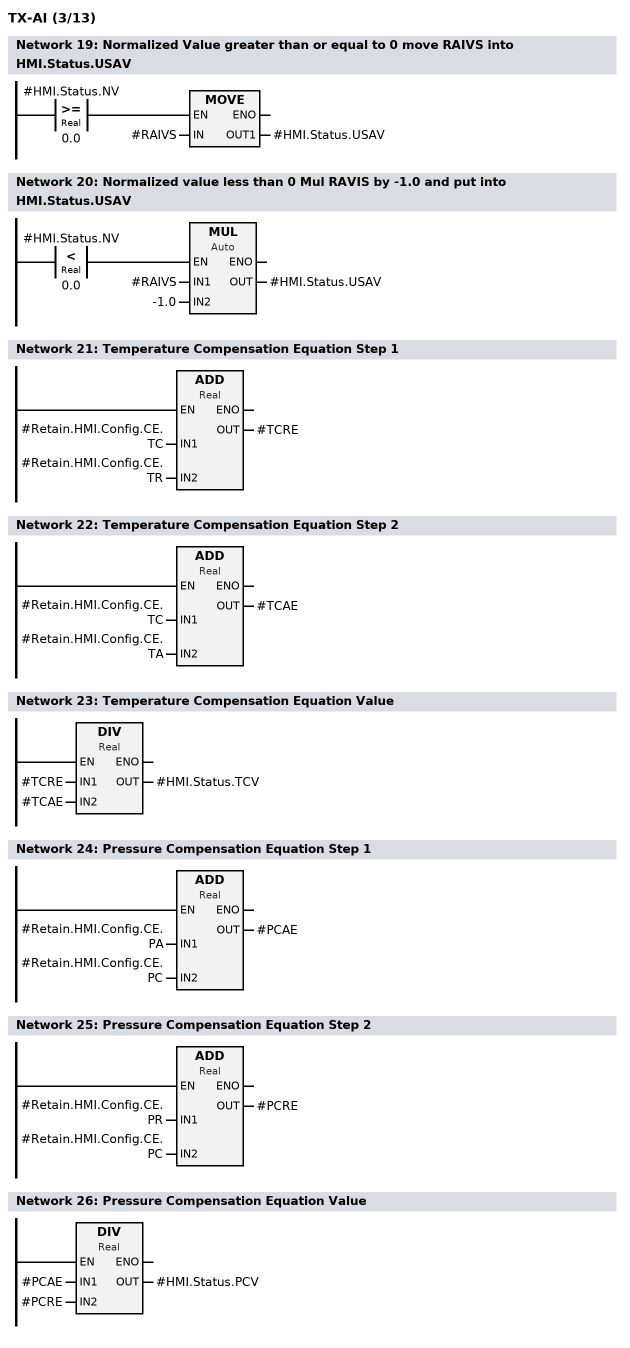
   RUNG wire#powerrail
      { S7_Templates := "SrcType := Real" } GE_Contact(in1 := #HMI.Status.NV, in2 := 0.0)
      { S7_GenerateENO := "TRUE" } Move(in := #RAIVS, out1 => #HMI.Status.USAV)
   END_RUNG
   // the same network as SCL:
   IF #HMI.Status.NV >= 0.0 THEN #HMI.Status.USAV := #RAIVS; END_IF;
END_REGION

REGION Network 20: Normalized value less than 0 Mul RAVIS by -1.0 and put into HMI.Status.USAV
   RUNG wire#powerrail
      { S7_Templates := "SrcType := Real" } LT_Contact(in1 := #HMI.Status.NV, in2 := 0.0)
      { S7_GenerateENO := "TRUE" } Mul(in1 := #RAIVS, in2 := -1.0, out => #HMI.Status.USAV)
   END_RUNG
   // the same network as SCL:
   IF #HMI.Status.NV < 0.0 THEN #HMI.Status.USAV := #RAIVS * (-1.0); END_IF;
END_REGION

REGION Network 21: Temperature Compensation Equation Step 1
   RUNG wire#powerrail
      { S7_Templates := "SrcType := Real"; S7_GenerateENO := "TRUE" } Add(in1 := #Retain.HMI.Config.CE.TC, in2 := #Retain.HMI.Config.CE.TR, out => #TCRE)
   END_RUNG
   // the same network as SCL:
   #TCRE := #Retain.HMI.Config.CE.TC + #Retain.HMI.Config.CE.TR;
END_REGION

REGION Network 22: Temperature Compensation Equation Step 2
   RUNG wire#powerrail
      { S7_Templates := "SrcType := Real"; S7_GenerateENO := "TRUE" } Add(in1 := #Retain.HMI.Config.CE.TC, in2 := #Retain.HMI.Config.CE.TA, out => #TCAE)
   END_RUNG
   // the same network as SCL:
   #TCAE := #Retain.HMI.Config.CE.TC + #Retain.HMI.Config.CE.TA;
END_REGION

REGION Network 23: Temperature Compensation Equation Value
   RUNG wire#powerrail
      { S7_Templates := "SrcType := Real"; S7_GenerateENO := "TRUE" } Div(in1 := #TCRE, in2 := #TCAE, out => #HMI.Status.TCV)
   END_RUNG
   // the same network as SCL:
   #HMI.Status.TCV := #TCRE / #TCAE;
END_REGION

REGION Network 24: Pressure Compensation Equation Step 1
   RUNG wire#powerrail
      { S7_Templates := "SrcType := Real"; S7_GenerateENO := "TRUE" } Add(in1 := #Retain.HMI.Config.CE.PA, in2 := #Retain.HMI.Config.CE.PC, out => #PCAE)
   END_RUNG
   // the same network as SCL:
   #PCAE := #Retain.HMI.Config.CE.PA + #Retain.HMI.Config.CE.PC;
END_REGION

REGION Network 25: Pressure Compensation Equation Step 2
   RUNG wire#powerrail
      { S7_Templates := "SrcType := Real"; S7_GenerateENO := "TRUE" } Add(in1 := #Retain.HMI.Config.CE.PR, in2 := #Retain.HMI.Config.CE.PC, out => #PCRE)
   END_RUNG
   // the same network as SCL:
   #PCRE := #Retain.HMI.Config.CE.PR + #Retain.HMI.Config.CE.PC;
END_REGION

REGION Network 26: Pressure Compensation Equation Value
   RUNG wire#powerrail
      { S7_Templates := "SrcType := Real"; S7_GenerateENO := "TRUE" } Div(in1 := #PCAE, in2 := #PCRE, out => #HMI.Status.PCV)
   END_RUNG
   // the same network as SCL:
   #HMI.Status.PCV := #PCAE / #PCRE;
END_REGION

REGION Network 27: Mol Weight Ratio
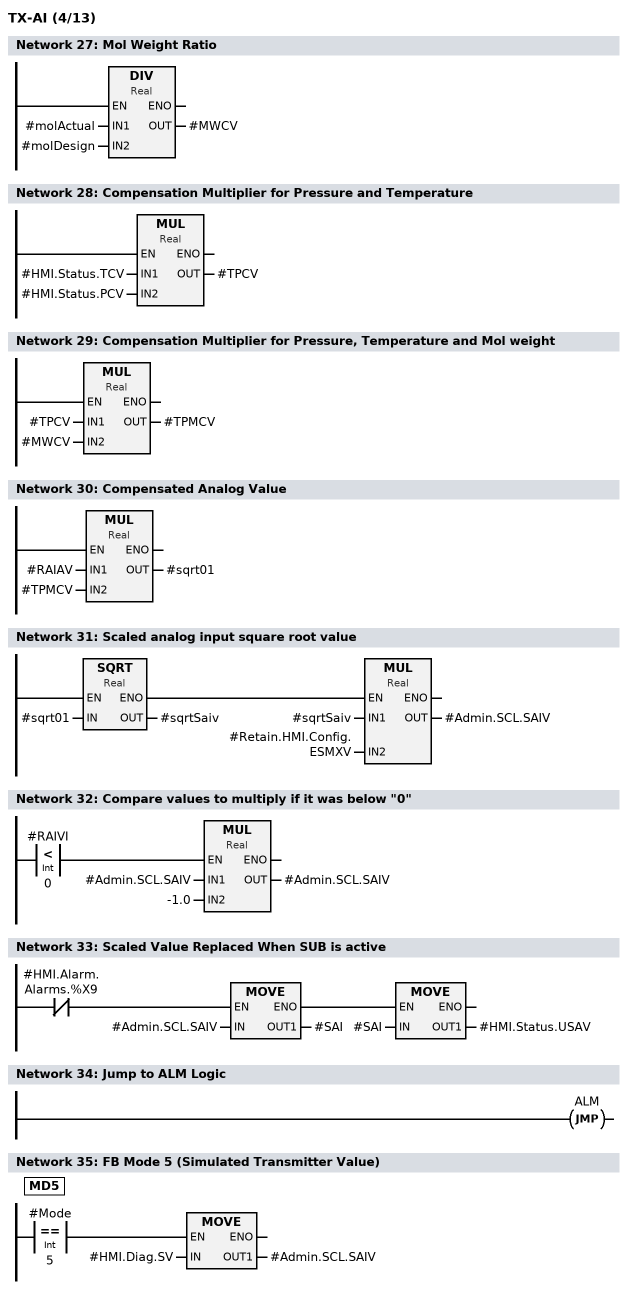
   RUNG wire#powerrail
      { S7_Templates := "SrcType := Real"; S7_GenerateENO := "TRUE" } Div(in1 := #molActual, in2 := #molDesign, out => #MWCV)
   END_RUNG
   // the same network as SCL:
   #MWCV := #molActual / #molDesign;
END_REGION

REGION Network 28: Compensation Multiplier for Pressure and Temperature
   RUNG wire#powerrail
      { S7_Templates := "SrcType := Real"; S7_GenerateENO := "TRUE" } Mul(in1 := #HMI.Status.TCV, in2 := #HMI.Status.PCV, out => #TPCV)
   END_RUNG
   // the same network as SCL:
   #TPCV := #HMI.Status.TCV * #HMI.Status.PCV;
END_REGION

REGION Network 29: Compensation Multiplier for Pressure, Temperature and Mol weight
   RUNG wire#powerrail
      { S7_Templates := "SrcType := Real"; S7_GenerateENO := "TRUE" } Mul(in1 := #TPCV, in2 := #MWCV, out => #TPMCV)
   END_RUNG
   // the same network as SCL:
   #TPMCV := #TPCV * #MWCV;
END_REGION

REGION Network 30: Compensated Analog Value
   RUNG wire#powerrail
      { S7_Templates := "SrcType := Real"; S7_GenerateENO := "TRUE" } Mul(in1 := #RAIAV, in2 := #TPMCV, out => #sqrt01)
   END_RUNG
   // the same network as SCL:
   #sqrt01 := #RAIAV * #TPMCV;
END_REGION

REGION Network 31: Scaled analog input square root value
   // ENO of a box is taken as its EN; it also drops when the box reports an error
   #sqrtSaiv := SQRT(#sqrt01);
   #Admin.SCL.SAIV := #sqrtSaiv * #Retain.HMI.Config.ESMXV;
END_REGION

REGION Network 32: Compare values to multiply if it was below "0"
   RUNG wire#powerrail
      { S7_Templates := "SrcType := Int" } LT_Contact(in1 := #RAIVI, in2 := 0)
      { S7_Templates := "SrcType := Real"; S7_GenerateENO := "TRUE" } Mul(in1 := #Admin.SCL.SAIV, in2 := -1.0, out => #Admin.SCL.SAIV)
   END_RUNG
   // the same network as SCL:
   IF #RAIVI < 0 THEN #Admin.SCL.SAIV := #Admin.SCL.SAIV * (-1.0); END_IF;
END_REGION

REGION Network 33: Scaled Value Replaced When SUB is active
   RUNG wire#powerrail
      I_Contact( #HMI.Alarm.Alarms.%X9 )
      { S7_GenerateENO := "TRUE" } Move(in := #Admin.SCL.SAIV, out1 => #SAI)
      { S7_GenerateENO := "TRUE" } Move(in := #SAI, out1 => #HMI.Status.USAV)
   END_RUNG
   // the same network as SCL:
   // ENO of a box is taken as its EN; it also drops when the box reports an error
   IF NOT #HMI.Alarm.Alarms.%X9 THEN
       #SAI := #Admin.SCL.SAIV;
       #HMI.Status.USAV := #SAI;
   END_IF;
END_REGION

REGION Network 34: Jump to ALM Logic
   RUNG wire#powerrail
      JumpCoil( ALM )
   END_RUNG
   // the same network as SCL:
   GOTO ALM;
END_REGION

REGION Network 35: FB Mode 5 (Simulated Transmitter Value)
   Label( MD5 )
   RUNG wire#powerrail
      { S7_Templates := "SrcType := Int" } EQ_Contact(in1 := #Mode, in2 := 5)
      { S7_GenerateENO := "TRUE" } Move(in := #HMI.Diag.SV, out1 => #Admin.SCL.SAIV)
   END_RUNG
   // the same network as SCL:
   MD5:
   IF #Mode = 5 THEN #Admin.SCL.SAIV := #HMI.Diag.SV; END_IF;
END_REGION

REGION Network 36: Scaled Value Replaced When SUB is active
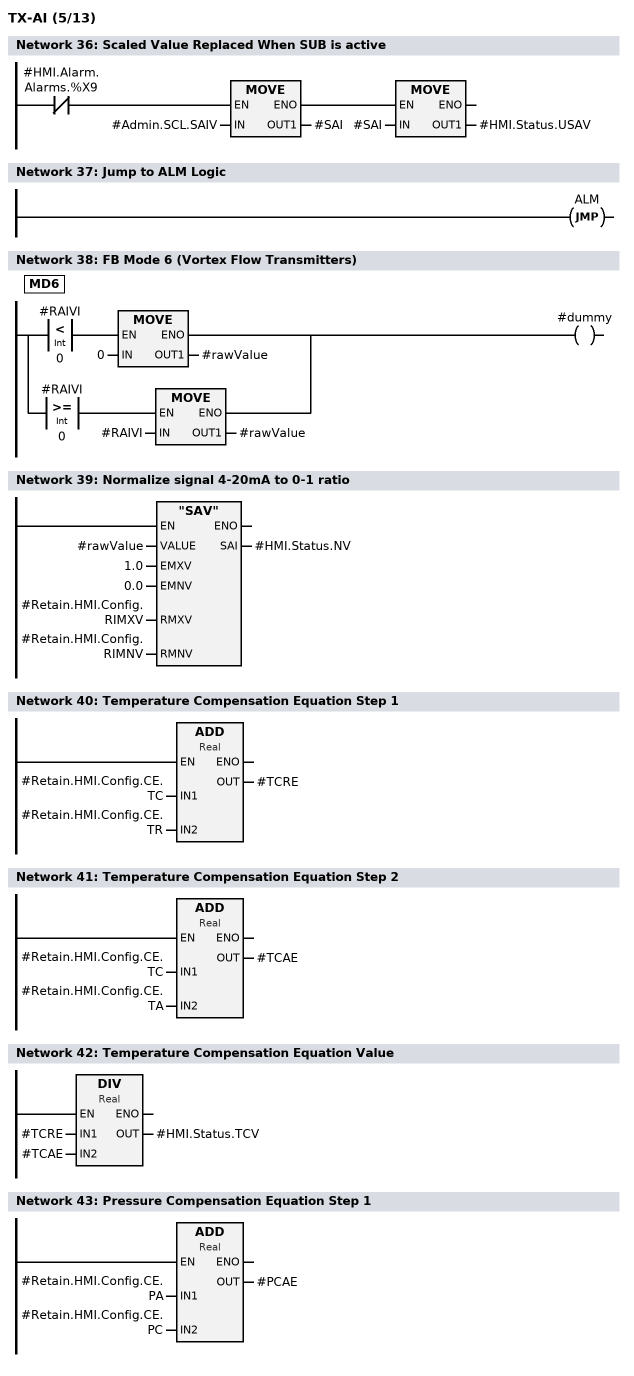
   RUNG wire#powerrail
      I_Contact( #HMI.Alarm.Alarms.%X9 )
      { S7_GenerateENO := "TRUE" } Move(in := #Admin.SCL.SAIV, out1 => #SAI)
      { S7_GenerateENO := "TRUE" } Move(in := #SAI, out1 => #HMI.Status.USAV)
   END_RUNG
   // the same network as SCL:
   // ENO of a box is taken as its EN; it also drops when the box reports an error
   IF NOT #HMI.Alarm.Alarms.%X9 THEN
       #SAI := #Admin.SCL.SAIV;
       #HMI.Status.USAV := #SAI;
   END_IF;
END_REGION

REGION Network 37: Jump to ALM Logic
   RUNG wire#powerrail
      JumpCoil( ALM )
   END_RUNG
   // the same network as SCL:
   GOTO ALM;
END_REGION

REGION Network 38: FB Mode 6 (Vortex Flow Transmitters)
   Label( MD6 )
   RUNG wire#powerrail
      { S7_Templates := "SrcType := Int" } LT_Contact(in1 := #RAIVI, in2 := 0)
      { S7_GenerateENO := "TRUE" } Move(in := 0, out1 => #rawValue)
      wire#w1
      Coil( #dummy )
   END_RUNG
   RUNG wire#powerrail
      { S7_Templates := "SrcType := Int" } GE_Contact(in1 := #RAIVI, in2 := 0)
      { S7_GenerateENO := "TRUE" } Move(in := #RAIVI, out1 => #rawValue)
   END_RUNG wire#w1
   // the same network as SCL:
   // ENO of a box is taken as its EN; it also drops when the box reports an error
   MD6:
   #_w1 := #RAIVI < 0;
   IF #_w1 THEN #rawValue := 0; END_IF;
   #_w2 := #RAIVI >= 0;
   IF #_w2 THEN #rawValue := #RAIVI; END_IF;
   #dummy := #_w1 OR #_w2;
END_REGION

REGION Network 39: Normalize signal 4-20mA to 0-1 ratio
   RUNG wire#powerrail
      "SAV"(VALUE := #rawValue, EMXV := 1.0, EMNV := 0.0, RMXV := #Retain.HMI.Config.RIMXV, RMNV := #Retain.HMI.Config.RIMNV, SAI => #HMI.Status.NV)
   END_RUNG
   // the same network as SCL:
   "SAV"(VALUE := #rawValue,
         EMXV := 1.0,
         EMNV := 0.0,
         RMXV := #Retain.HMI.Config.RIMXV,
         RMNV := #Retain.HMI.Config.RIMNV,
         SAI => #HMI.Status.NV);
END_REGION

REGION Network 40: Temperature Compensation Equation Step 1
   RUNG wire#powerrail
      { S7_Templates := "SrcType := Real"; S7_GenerateENO := "TRUE" } Add(in1 := #Retain.HMI.Config.CE.TC, in2 := #Retain.HMI.Config.CE.TR, out => #TCRE)
   END_RUNG
   // the same network as SCL:
   #TCRE := #Retain.HMI.Config.CE.TC + #Retain.HMI.Config.CE.TR;
END_REGION

REGION Network 41: Temperature Compensation Equation Step 2
   RUNG wire#powerrail
      { S7_Templates := "SrcType := Real"; S7_GenerateENO := "TRUE" } Add(in1 := #Retain.HMI.Config.CE.TC, in2 := #Retain.HMI.Config.CE.TA, out => #TCAE)
   END_RUNG
   // the same network as SCL:
   #TCAE := #Retain.HMI.Config.CE.TC + #Retain.HMI.Config.CE.TA;
END_REGION

REGION Network 42: Temperature Compensation Equation Value
   RUNG wire#powerrail
      { S7_Templates := "SrcType := Real"; S7_GenerateENO := "TRUE" } Div(in1 := #TCRE, in2 := #TCAE, out => #HMI.Status.TCV)
   END_RUNG
   // the same network as SCL:
   #HMI.Status.TCV := #TCRE / #TCAE;
END_REGION

REGION Network 43: Pressure Compensation Equation Step 1
   RUNG wire#powerrail
      { S7_Templates := "SrcType := Real"; S7_GenerateENO := "TRUE" } Add(in1 := #Retain.HMI.Config.CE.PA, in2 := #Retain.HMI.Config.CE.PC, out => #PCAE)
   END_RUNG
   // the same network as SCL:
   #PCAE := #Retain.HMI.Config.CE.PA + #Retain.HMI.Config.CE.PC;
END_REGION

REGION Network 44: Pressure Compensation Equation Step 2
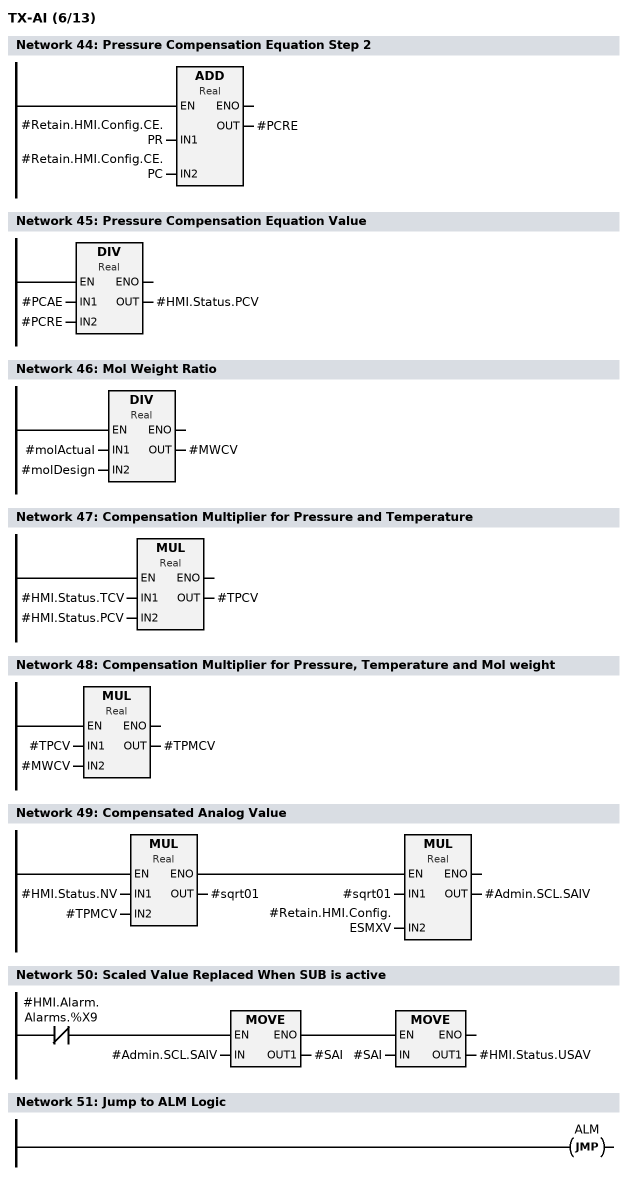
   RUNG wire#powerrail
      { S7_Templates := "SrcType := Real"; S7_GenerateENO := "TRUE" } Add(in1 := #Retain.HMI.Config.CE.PR, in2 := #Retain.HMI.Config.CE.PC, out => #PCRE)
   END_RUNG
   // the same network as SCL:
   #PCRE := #Retain.HMI.Config.CE.PR + #Retain.HMI.Config.CE.PC;
END_REGION

REGION Network 45: Pressure Compensation Equation Value
   RUNG wire#powerrail
      { S7_Templates := "SrcType := Real"; S7_GenerateENO := "TRUE" } Div(in1 := #PCAE, in2 := #PCRE, out => #HMI.Status.PCV)
   END_RUNG
   // the same network as SCL:
   #HMI.Status.PCV := #PCAE / #PCRE;
END_REGION

REGION Network 46: Mol Weight Ratio
   RUNG wire#powerrail
      { S7_Templates := "SrcType := Real"; S7_GenerateENO := "TRUE" } Div(in1 := #molActual, in2 := #molDesign, out => #MWCV)
   END_RUNG
   // the same network as SCL:
   #MWCV := #molActual / #molDesign;
END_REGION

REGION Network 47: Compensation Multiplier for Pressure and Temperature
   RUNG wire#powerrail
      { S7_Templates := "SrcType := Real"; S7_GenerateENO := "TRUE" } Mul(in1 := #HMI.Status.TCV, in2 := #HMI.Status.PCV, out => #TPCV)
   END_RUNG
   // the same network as SCL:
   #TPCV := #HMI.Status.TCV * #HMI.Status.PCV;
END_REGION

REGION Network 48: Compensation Multiplier for Pressure, Temperature and Mol weight
   RUNG wire#powerrail
      { S7_Templates := "SrcType := Real"; S7_GenerateENO := "TRUE" } Mul(in1 := #TPCV, in2 := #MWCV, out => #TPMCV)
   END_RUNG
   // the same network as SCL:
   #TPMCV := #TPCV * #MWCV;
END_REGION

REGION Network 49: Compensated Analog Value
   RUNG wire#powerrail
      { S7_Templates := "SrcType := Real"; S7_GenerateENO := "TRUE" } Mul(in1 := #HMI.Status.NV, in2 := #TPMCV, out => #sqrt01)
      { S7_Templates := "SrcType := Real"; S7_GenerateENO := "TRUE" } Mul(in1 := #sqrt01, in2 := #Retain.HMI.Config.ESMXV, out => #Admin.SCL.SAIV)
   END_RUNG
   // the same network as SCL:
   // ENO of a box is taken as its EN; it also drops when the box reports an error
   #sqrt01 := #HMI.Status.NV * #TPMCV;
   #Admin.SCL.SAIV := #sqrt01 * #Retain.HMI.Config.ESMXV;
END_REGION

REGION Network 50: Scaled Value Replaced When SUB is active
   RUNG wire#powerrail
      I_Contact( #HMI.Alarm.Alarms.%X9 )
      { S7_GenerateENO := "TRUE" } Move(in := #Admin.SCL.SAIV, out1 => #SAI)
      { S7_GenerateENO := "TRUE" } Move(in := #SAI, out1 => #HMI.Status.USAV)
   END_RUNG
   // the same network as SCL:
   // ENO of a box is taken as its EN; it also drops when the box reports an error
   IF NOT #HMI.Alarm.Alarms.%X9 THEN
       #SAI := #Admin.SCL.SAIV;
       #HMI.Status.USAV := #SAI;
   END_IF;
END_REGION

REGION Network 51: Jump to ALM Logic
   RUNG wire#powerrail
      JumpCoil( ALM )
   END_RUNG
   // the same network as SCL:
   GOTO ALM;
END_REGION

REGION Network 52: ALM (Global Hold Preset Time Condition)
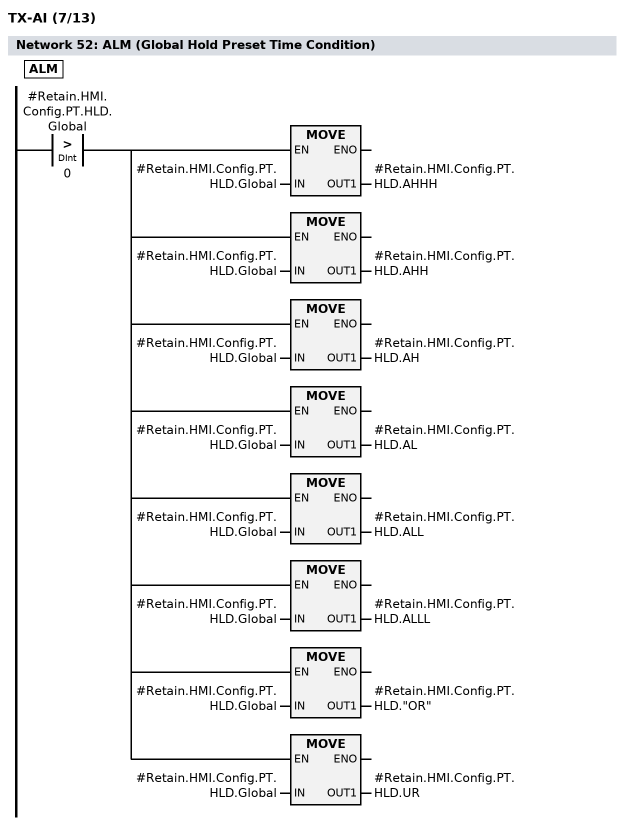
   Label( ALM )
   RUNG wire#powerrail
      { S7_Templates := "SrcType := DInt" } GT_Contact(in1 := #Retain.HMI.Config.PT.HLD.Global, in2 := 0)
      wire#w1
      { S7_GenerateENO := "TRUE" } Move(in := #Retain.HMI.Config.PT.HLD.Global, out1 => #Retain.HMI.Config.PT.HLD.AHHH)
   END_RUNG
   RUNG wire#w1
      { S7_GenerateENO := "TRUE" } Move(in := #Retain.HMI.Config.PT.HLD.Global, out1 => #Retain.HMI.Config.PT.HLD.AHH)
   END_RUNG
   RUNG wire#w1
      { S7_GenerateENO := "TRUE" } Move(in := #Retain.HMI.Config.PT.HLD.Global, out1 => #Retain.HMI.Config.PT.HLD.AH)
   END_RUNG
   RUNG wire#w1
      { S7_GenerateENO := "TRUE" } Move(in := #Retain.HMI.Config.PT.HLD.Global, out1 => #Retain.HMI.Config.PT.HLD.AL)
   END_RUNG
   RUNG wire#w1
      { S7_GenerateENO := "TRUE" } Move(in := #Retain.HMI.Config.PT.HLD.Global, out1 => #Retain.HMI.Config.PT.HLD.ALL)
   END_RUNG
   RUNG wire#w1
      { S7_GenerateENO := "TRUE" } Move(in := #Retain.HMI.Config.PT.HLD.Global, out1 => #Retain.HMI.Config.PT.HLD.ALLL)
   END_RUNG
   RUNG wire#w1
      { S7_GenerateENO := "TRUE" } Move(in := #Retain.HMI.Config.PT.HLD.Global, out1 => #Retain.HMI.Config.PT.HLD."OR")
   END_RUNG
   RUNG wire#w1
      { S7_GenerateENO := "TRUE" } Move(in := #Retain.HMI.Config.PT.HLD.Global, out1 => #Retain.HMI.Config.PT.HLD.UR)
   END_RUNG
   // the same network as SCL:
   ALM:
   IF #Retain.HMI.Config.PT.HLD.Global > 0 THEN
       #Retain.HMI.Config.PT.HLD.AHHH := #Retain.HMI.Config.PT.HLD.Global;
       #Retain.HMI.Config.PT.HLD.AHH := #Retain.HMI.Config.PT.HLD.Global;
       #Retain.HMI.Config.PT.HLD.AH := #Retain.HMI.Config.PT.HLD.Global;
       #Retain.HMI.Config.PT.HLD.AL := #Retain.HMI.Config.PT.HLD.Global;
       #Retain.HMI.Config.PT.HLD.ALL := #Retain.HMI.Config.PT.HLD.Global;
       #Retain.HMI.Config.PT.HLD.ALLL := #Retain.HMI.Config.PT.HLD.Global;
       #Retain.HMI.Config.PT.HLD."OR" := #Retain.HMI.Config.PT.HLD.Global;
       #Retain.HMI.Config.PT.HLD.UR := #Retain.HMI.Config.PT.HLD.Global;
   END_IF;
END_REGION

REGION Network 53: Global Debounce Preset Time Condition
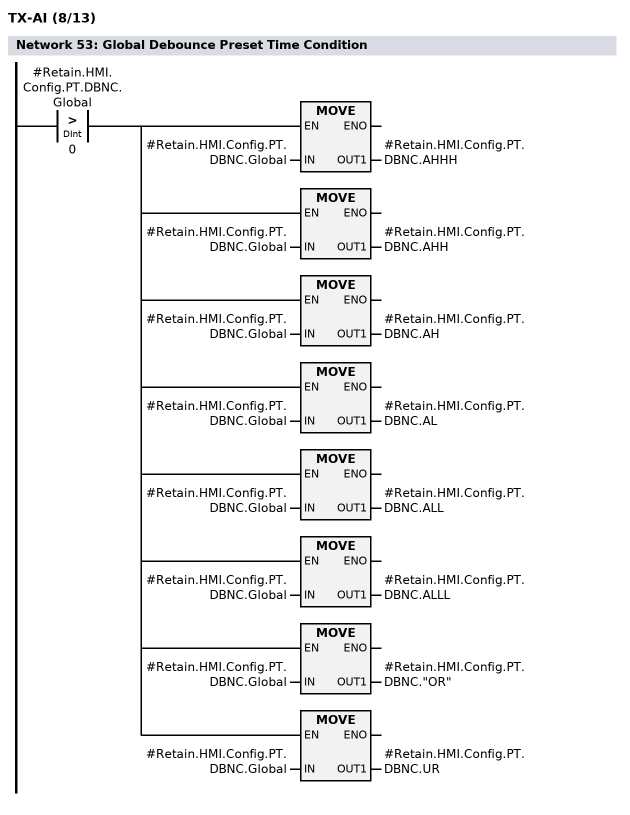
   RUNG wire#powerrail
      { S7_Templates := "SrcType := DInt" } GT_Contact(in1 := #Retain.HMI.Config.PT.DBNC.Global, in2 := 0)
      wire#w1
      { S7_GenerateENO := "TRUE" } Move(in := #Retain.HMI.Config.PT.DBNC.Global, out1 => #Retain.HMI.Config.PT.DBNC.AHHH)
   END_RUNG
   RUNG wire#w1
      { S7_GenerateENO := "TRUE" } Move(in := #Retain.HMI.Config.PT.DBNC.Global, out1 => #Retain.HMI.Config.PT.DBNC.AHH)
   END_RUNG
   RUNG wire#w1
      { S7_GenerateENO := "TRUE" } Move(in := #Retain.HMI.Config.PT.DBNC.Global, out1 => #Retain.HMI.Config.PT.DBNC.AH)
   END_RUNG
   RUNG wire#w1
      { S7_GenerateENO := "TRUE" } Move(in := #Retain.HMI.Config.PT.DBNC.Global, out1 => #Retain.HMI.Config.PT.DBNC.AL)
   END_RUNG
   RUNG wire#w1
      { S7_GenerateENO := "TRUE" } Move(in := #Retain.HMI.Config.PT.DBNC.Global, out1 => #Retain.HMI.Config.PT.DBNC.ALL)
   END_RUNG
   RUNG wire#w1
      { S7_GenerateENO := "TRUE" } Move(in := #Retain.HMI.Config.PT.DBNC.Global, out1 => #Retain.HMI.Config.PT.DBNC.ALLL)
   END_RUNG
   RUNG wire#w1
      { S7_GenerateENO := "TRUE" } Move(in := #Retain.HMI.Config.PT.DBNC.Global, out1 => #Retain.HMI.Config.PT.DBNC."OR")
   END_RUNG
   RUNG wire#w1
      { S7_GenerateENO := "TRUE" } Move(in := #Retain.HMI.Config.PT.DBNC.Global, out1 => #Retain.HMI.Config.PT.DBNC.UR)
   END_RUNG
   // the same network as SCL:
   IF #Retain.HMI.Config.PT.DBNC.Global > 0 THEN
       #Retain.HMI.Config.PT.DBNC.AHHH := #Retain.HMI.Config.PT.DBNC.Global;
       #Retain.HMI.Config.PT.DBNC.AHH := #Retain.HMI.Config.PT.DBNC.Global;
       #Retain.HMI.Config.PT.DBNC.AH := #Retain.HMI.Config.PT.DBNC.Global;
       #Retain.HMI.Config.PT.DBNC.AL := #Retain.HMI.Config.PT.DBNC.Global;
       #Retain.HMI.Config.PT.DBNC.ALL := #Retain.HMI.Config.PT.DBNC.Global;
       #Retain.HMI.Config.PT.DBNC.ALLL := #Retain.HMI.Config.PT.DBNC.Global;
       #Retain.HMI.Config.PT.DBNC."OR" := #Retain.HMI.Config.PT.DBNC.Global;
       #Retain.HMI.Config.PT.DBNC.UR := #Retain.HMI.Config.PT.DBNC.Global;
   END_IF;
END_REGION

REGION Network 54: Global Hysteresis Setpoint Condition
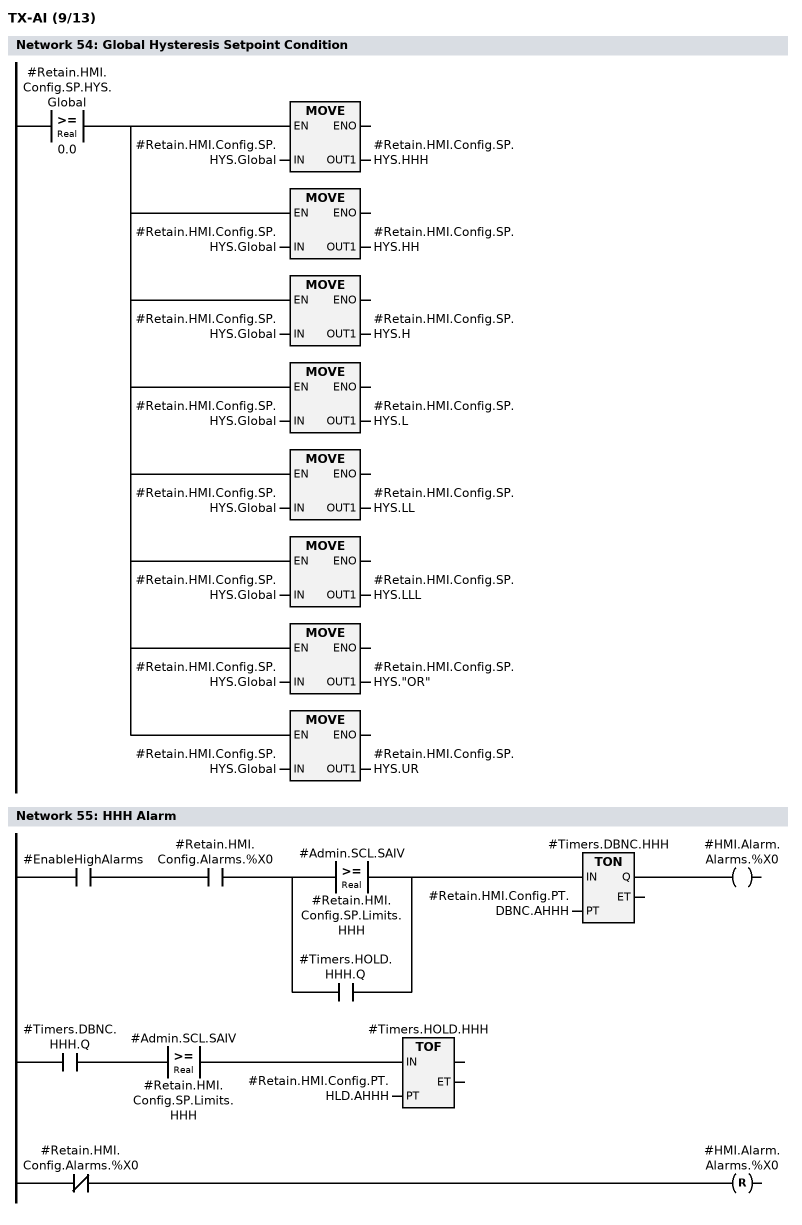
   RUNG wire#powerrail
      { S7_Templates := "SrcType := Real" } GE_Contact(in1 := #Retain.HMI.Config.SP.HYS.Global, in2 := 0.0)
      wire#w1
      { S7_GenerateENO := "TRUE" } Move(in := #Retain.HMI.Config.SP.HYS.Global, out1 => #Retain.HMI.Config.SP.HYS.HHH)
   END_RUNG
   RUNG wire#w1
      { S7_GenerateENO := "TRUE" } Move(in := #Retain.HMI.Config.SP.HYS.Global, out1 => #Retain.HMI.Config.SP.HYS.HH)
   END_RUNG
   RUNG wire#w1
      { S7_GenerateENO := "TRUE" } Move(in := #Retain.HMI.Config.SP.HYS.Global, out1 => #Retain.HMI.Config.SP.HYS.H)
   END_RUNG
   RUNG wire#w1
      { S7_GenerateENO := "TRUE" } Move(in := #Retain.HMI.Config.SP.HYS.Global, out1 => #Retain.HMI.Config.SP.HYS.L)
   END_RUNG
   RUNG wire#w1
      { S7_GenerateENO := "TRUE" } Move(in := #Retain.HMI.Config.SP.HYS.Global, out1 => #Retain.HMI.Config.SP.HYS.LL)
   END_RUNG
   RUNG wire#w1
      { S7_GenerateENO := "TRUE" } Move(in := #Retain.HMI.Config.SP.HYS.Global, out1 => #Retain.HMI.Config.SP.HYS.LLL)
   END_RUNG
   RUNG wire#w1
      { S7_GenerateENO := "TRUE" } Move(in := #Retain.HMI.Config.SP.HYS.Global, out1 => #Retain.HMI.Config.SP.HYS."OR")
   END_RUNG
   RUNG wire#w1
      { S7_GenerateENO := "TRUE" } Move(in := #Retain.HMI.Config.SP.HYS.Global, out1 => #Retain.HMI.Config.SP.HYS.UR)
   END_RUNG
   // the same network as SCL:
   IF #Retain.HMI.Config.SP.HYS.Global >= 0.0 THEN
       #Retain.HMI.Config.SP.HYS.HHH := #Retain.HMI.Config.SP.HYS.Global;
       #Retain.HMI.Config.SP.HYS.HH := #Retain.HMI.Config.SP.HYS.Global;
       #Retain.HMI.Config.SP.HYS.H := #Retain.HMI.Config.SP.HYS.Global;
       #Retain.HMI.Config.SP.HYS.L := #Retain.HMI.Config.SP.HYS.Global;
       #Retain.HMI.Config.SP.HYS.LL := #Retain.HMI.Config.SP.HYS.Global;
       #Retain.HMI.Config.SP.HYS.LLL := #Retain.HMI.Config.SP.HYS.Global;
       #Retain.HMI.Config.SP.HYS."OR" := #Retain.HMI.Config.SP.HYS.Global;
       #Retain.HMI.Config.SP.HYS.UR := #Retain.HMI.Config.SP.HYS.Global;
   END_IF;
END_REGION

REGION Network 55: HHH Alarm
   #Timers.DBNC.HHH.TON(IN := #EnableHighAlarms AND #Retain.HMI.Config.Alarms.%X0 AND ((#Admin.SCL.SAIV >= #Retain.HMI.Config.SP.Limits.HHH) OR #Timers.HOLD.HHH.Q),
                        PT := #Retain.HMI.Config.PT.DBNC.AHHH);
   #HMI.Alarm.Alarms.%X0 := #Timers.DBNC.HHH.Q;
   #Timers.HOLD.HHH.TOF(IN := #Timers.DBNC.HHH.Q AND (#Admin.SCL.SAIV >= #Retain.HMI.Config.SP.Limits.HHH),
                        PT := #Retain.HMI.Config.PT.HLD.AHHH);
   IF NOT #Retain.HMI.Config.Alarms.%X0 THEN #HMI.Alarm.Alarms.%X0 := FALSE; END_IF;
END_REGION

REGION Network 56: HH Alarm
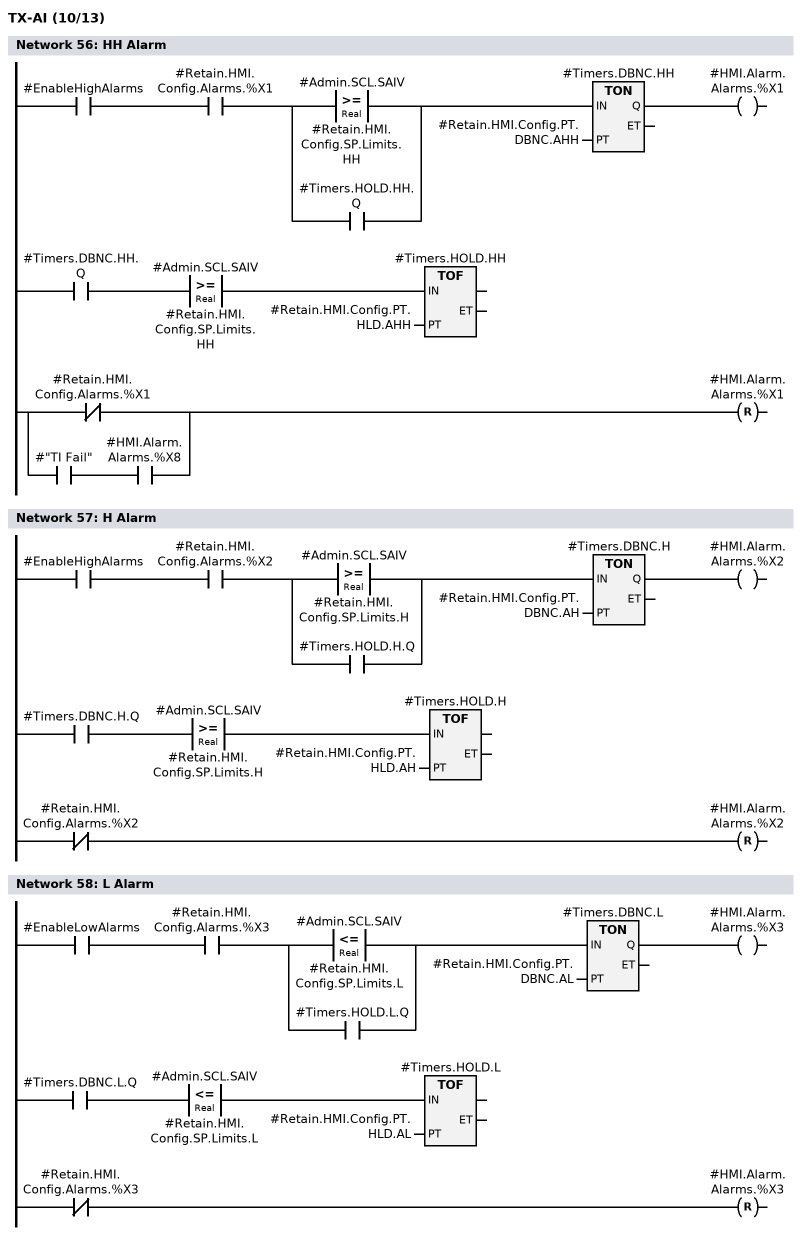
   #Timers.DBNC.HH.TON(IN := #EnableHighAlarms AND #Retain.HMI.Config.Alarms.%X1 AND ((#Admin.SCL.SAIV >= #Retain.HMI.Config.SP.Limits.HH) OR #Timers.HOLD.HH.Q),
                       PT := #Retain.HMI.Config.PT.DBNC.AHH);
   #HMI.Alarm.Alarms.%X1 := #Timers.DBNC.HH.Q;
   #Timers.HOLD.HH.TOF(IN := #Timers.DBNC.HH.Q AND (#Admin.SCL.SAIV >= #Retain.HMI.Config.SP.Limits.HH),
                       PT := #Retain.HMI.Config.PT.HLD.AHH);
   IF NOT #Retain.HMI.Config.Alarms.%X1 OR (#"TI Fail" AND #HMI.Alarm.Alarms.%X8) THEN
       #HMI.Alarm.Alarms.%X1 := FALSE;
   END_IF;
END_REGION

REGION Network 57: H Alarm
   #Timers.DBNC.H.TON(IN := #EnableHighAlarms AND #Retain.HMI.Config.Alarms.%X2 AND ((#Admin.SCL.SAIV >= #Retain.HMI.Config.SP.Limits.H) OR #Timers.HOLD.H.Q),
                      PT := #Retain.HMI.Config.PT.DBNC.AH);
   #HMI.Alarm.Alarms.%X2 := #Timers.DBNC.H.Q;
   #Timers.HOLD.H.TOF(IN := #Timers.DBNC.H.Q AND (#Admin.SCL.SAIV >= #Retain.HMI.Config.SP.Limits.H),
                      PT := #Retain.HMI.Config.PT.HLD.AH);
   IF NOT #Retain.HMI.Config.Alarms.%X2 THEN #HMI.Alarm.Alarms.%X2 := FALSE; END_IF;
END_REGION

REGION Network 58: L Alarm
   #Timers.DBNC.L.TON(IN := #EnableLowAlarms AND #Retain.HMI.Config.Alarms.%X3 AND ((#Admin.SCL.SAIV <= #Retain.HMI.Config.SP.Limits.L) OR #Timers.HOLD.L.Q),
                      PT := #Retain.HMI.Config.PT.DBNC.AL);
   #HMI.Alarm.Alarms.%X3 := #Timers.DBNC.L.Q;
   #Timers.HOLD.L.TOF(IN := #Timers.DBNC.L.Q AND (#Admin.SCL.SAIV <= #Retain.HMI.Config.SP.Limits.L),
                      PT := #Retain.HMI.Config.PT.HLD.AL);
   IF NOT #Retain.HMI.Config.Alarms.%X3 THEN #HMI.Alarm.Alarms.%X3 := FALSE; END_IF;
END_REGION

REGION Network 59: LL Alarm
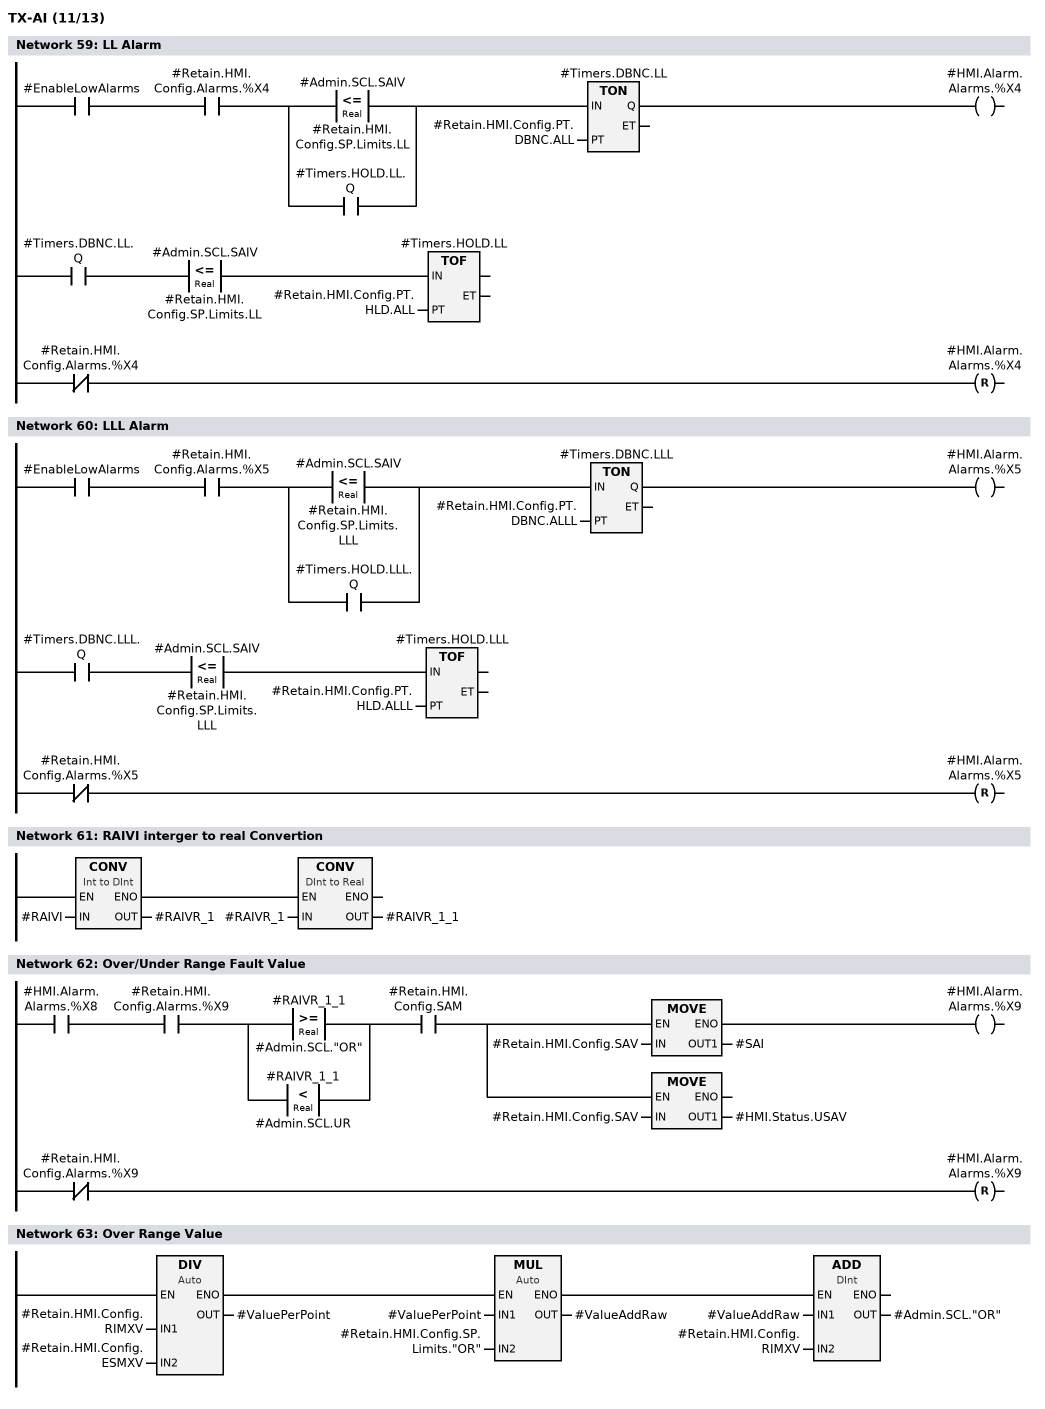
   #Timers.DBNC.LL.TON(IN := #EnableLowAlarms AND #Retain.HMI.Config.Alarms.%X4 AND ((#Admin.SCL.SAIV <= #Retain.HMI.Config.SP.Limits.LL) OR #Timers.HOLD.LL.Q),
                       PT := #Retain.HMI.Config.PT.DBNC.ALL);
   #HMI.Alarm.Alarms.%X4 := #Timers.DBNC.LL.Q;
   #Timers.HOLD.LL.TOF(IN := #Timers.DBNC.LL.Q AND (#Admin.SCL.SAIV <= #Retain.HMI.Config.SP.Limits.LL),
                       PT := #Retain.HMI.Config.PT.HLD.ALL);
   IF NOT #Retain.HMI.Config.Alarms.%X4 THEN #HMI.Alarm.Alarms.%X4 := FALSE; END_IF;
END_REGION

REGION Network 60: LLL Alarm
   #Timers.DBNC.LLL.TON(IN := #EnableLowAlarms AND #Retain.HMI.Config.Alarms.%X5 AND ((#Admin.SCL.SAIV <= #Retain.HMI.Config.SP.Limits.LLL) OR #Timers.HOLD.LLL.Q),
                        PT := #Retain.HMI.Config.PT.DBNC.ALLL);
   #HMI.Alarm.Alarms.%X5 := #Timers.DBNC.LLL.Q;
   #Timers.HOLD.LLL.TOF(IN := #Timers.DBNC.LLL.Q AND (#Admin.SCL.SAIV <= #Retain.HMI.Config.SP.Limits.LLL),
                        PT := #Retain.HMI.Config.PT.HLD.ALLL);
   IF NOT #Retain.HMI.Config.Alarms.%X5 THEN #HMI.Alarm.Alarms.%X5 := FALSE; END_IF;
END_REGION

REGION Network 61: RAIVI interger to real Convertion
   RUNG wire#powerrail
      { S7_Templates := "[SrcType := Int, DestType := DInt]"; S7_GenerateENO := "TRUE" } Convert(in := #RAIVI, out => #RAIVR_1)
      { S7_Templates := "[SrcType := DInt, DestType := Real]"; S7_GenerateENO := "TRUE" } Convert(in := #RAIVR_1, out => #RAIVR_1_1)
   END_RUNG
   // the same network as SCL:
   // ENO of a box is taken as its EN; it also drops when the box reports an error
   #RAIVR_1 := INT_TO_DINT(#RAIVI);
   #RAIVR_1_1 := DINT_TO_REAL(#RAIVR_1);
END_REGION

REGION Network 62: Over/Under Range Fault Value
   RUNG wire#powerrail
      Contact( #HMI.Alarm.Alarms.%X8 )
      Contact( #Retain.HMI.Config.Alarms.%X9 )
      wire#w1
      { S7_Templates := "SrcType := Real" } GE_Contact(in1 := #RAIVR_1_1, in2 := #Admin.SCL."OR")
      wire#w2
      Contact( #Retain.HMI.Config.SAM )
      wire#w3
      { S7_GenerateENO := "TRUE" } Move(in := #Retain.HMI.Config.SAV, out1 => #SAI)
      Coil( #HMI.Alarm.Alarms.%X9 )
   END_RUNG
   RUNG wire#w1
      { S7_Templates := "SrcType := Real" } LT_Contact(in1 := #RAIVR_1_1, in2 := #Admin.SCL.UR)
   END_RUNG wire#w2
   RUNG wire#w3
      { S7_GenerateENO := "TRUE" } Move(in := #Retain.HMI.Config.SAV, out1 => #HMI.Status.USAV)
   END_RUNG
   RUNG wire#powerrail
      I_Contact( #Retain.HMI.Config.Alarms.%X9 )
      R_Coil( #HMI.Alarm.Alarms.%X9 )
   END_RUNG
   // the same network as SCL:
   // ENO of a box is taken as its EN; it also drops when the box reports an error
   #_w1 := #HMI.Alarm.Alarms.%X8 AND #Retain.HMI.Config.Alarms.%X9 AND ((#RAIVR_1_1 >= #Admin.SCL."OR") OR (#RAIVR_1_1 < #Admin.SCL.UR)) AND #Retain.HMI.Config.SAM;
   IF #_w1 THEN #SAI := #Retain.HMI.Config.SAV; END_IF;
   #HMI.Alarm.Alarms.%X9 := #_w1;
   IF #_w1 THEN #HMI.Status.USAV := #Retain.HMI.Config.SAV; END_IF;
   IF NOT #Retain.HMI.Config.Alarms.%X9 THEN #HMI.Alarm.Alarms.%X9 := FALSE; END_IF;
END_REGION

REGION Network 63: Over Range Value
   RUNG wire#powerrail
      Div(in1 := #Retain.HMI.Config.RIMXV, in2 := #Retain.HMI.Config.ESMXV, out => #ValuePerPoint)
      Mul(in1 := #ValuePerPoint, in2 := #Retain.HMI.Config.SP.Limits."OR", out => #ValueAddRaw)
      { S7_Templates := "SrcType := DInt"; S7_GenerateENO := "TRUE" } Add(in1 := #ValueAddRaw, in2 := #Retain.HMI.Config.RIMXV, out => #Admin.SCL."OR")
   END_RUNG
   // the same network as SCL:
   #ValuePerPoint := #Retain.HMI.Config.RIMXV / #Retain.HMI.Config.ESMXV;
   #ValueAddRaw := #ValuePerPoint * #Retain.HMI.Config.SP.Limits."OR";
   #Admin.SCL."OR" := #ValueAddRaw + #Retain.HMI.Config.RIMXV;
END_REGION

REGION Network 64: Under Range Value
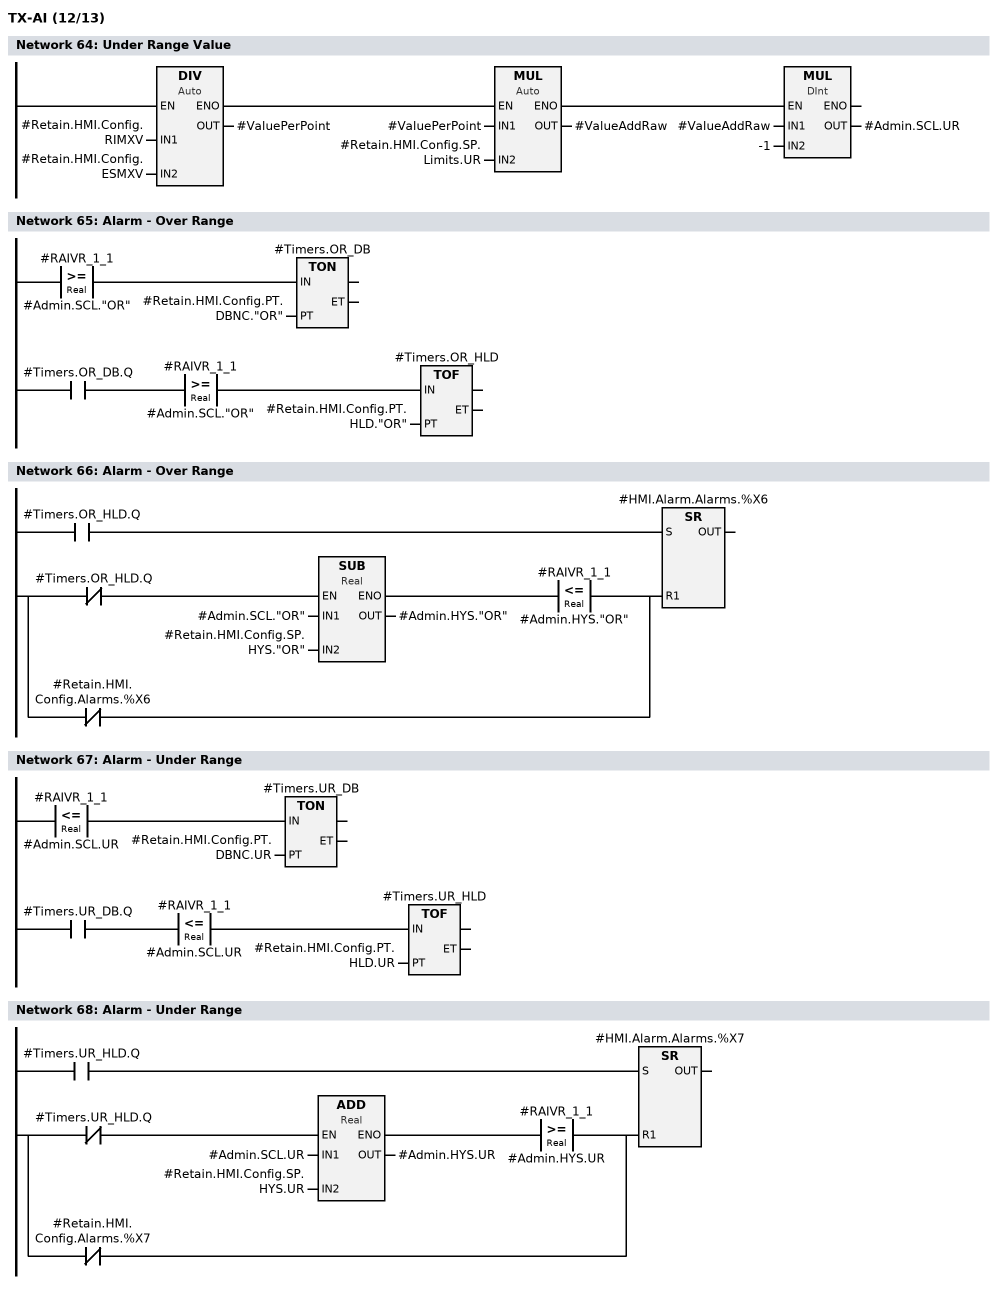
   RUNG wire#powerrail
      Div(in1 := #Retain.HMI.Config.RIMXV, in2 := #Retain.HMI.Config.ESMXV, out => #ValuePerPoint)
      Mul(in1 := #ValuePerPoint, in2 := #Retain.HMI.Config.SP.Limits.UR, out => #ValueAddRaw)
      { S7_Templates := "SrcType := DInt"; S7_GenerateENO := "TRUE" } Mul(in1 := #ValueAddRaw, in2 := -1, out => #Admin.SCL.UR)
   END_RUNG
   // the same network as SCL:
   #ValuePerPoint := #Retain.HMI.Config.RIMXV / #Retain.HMI.Config.ESMXV;
   #ValueAddRaw := #ValuePerPoint * #Retain.HMI.Config.SP.Limits.UR;
   #Admin.SCL.UR := #ValueAddRaw * (-1);
END_REGION

REGION Network 65: Alarm - Over Range
   #Timers.OR_DB.TON(IN := #RAIVR_1_1 >= #Admin.SCL."OR", PT := #Retain.HMI.Config.PT.DBNC."OR");
   #Timers.OR_HLD.TOF(IN := #Timers.OR_DB.Q AND (#RAIVR_1_1 >= #Admin.SCL."OR"),
                      PT := #Retain.HMI.Config.PT.HLD."OR");
END_REGION

REGION Network 66: Alarm - Over Range
   RUNG wire#powerrail
      Contact( #Timers.OR_HLD.Q )
      S_SR(operand := #HMI.Alarm.Alarms.%X6, r1 := wire#w1)
   END_RUNG
   RUNG wire#powerrail
      I_Contact( #Timers.OR_HLD.Q )
      { S7_Templates := "SrcType := Real"; S7_GenerateENO := "TRUE" } Sub(in1 := #Admin.SCL."OR", in2 := #Retain.HMI.Config.SP.HYS."OR", out => #Admin.HYS."OR")
      { S7_Templates := "SrcType := Real" } LE_Contact(in1 := #RAIVR_1_1, in2 := #Admin.HYS."OR")
   END_RUNG wire#w1
   RUNG wire#powerrail
      I_Contact( #Retain.HMI.Config.Alarms.%X6 )
   END_RUNG wire#w1
   // the same network as SCL:
   // ENO of a box is taken as its EN; it also drops when the box reports an error
   IF NOT #Timers.OR_HLD.Q THEN #Admin.HYS."OR" := #Admin.SCL."OR" - #Retain.HMI.Config.SP.HYS."OR"; END_IF;
   IF #Timers.OR_HLD.Q THEN
       #HMI.Alarm.Alarms.%X6 := TRUE;   // SR flip-flop
   END_IF;
   IF (NOT #Timers.OR_HLD.Q AND (#RAIVR_1_1 <= #Admin.HYS."OR")) OR NOT #Retain.HMI.Config.Alarms.%X6 THEN
       #HMI.Alarm.Alarms.%X6 := FALSE;
   END_IF;
END_REGION

REGION Network 67: Alarm - Under Range
   #Timers.UR_DB.TON(IN := #RAIVR_1_1 <= #Admin.SCL.UR, PT := #Retain.HMI.Config.PT.DBNC.UR);
   #Timers.UR_HLD.TOF(IN := #Timers.UR_DB.Q AND (#RAIVR_1_1 <= #Admin.SCL.UR),
                      PT := #Retain.HMI.Config.PT.HLD.UR);
END_REGION

